// Mitsubishi GX Works2 project: 30国轩预化成10.29   PLC: Q10UDEH (continued)

Rotor30403(ShuttleCarInOut:=RotorIO30403);(*预化成2入库转台*)
RotorIO30403.xReady:=XAD;
Y264:=RotorIO30403.xCW;					
Y265:=RotorIO30403.xCCW;	
Y285:=RotorIO30403.xBrake;				
RotorIO30403.xForward:=M545;					
RotorIO30403.xBackward:=M546;					
ShuttleCarCurrentPosition(X65 OR X64,X65,X64,FALSE,RotorIO30403.iCurrentPos);					
M647:=RotorIO30403.xOvertimeAlarm ;					
RotorIO30403.diDeviceID:=30403;					
RotorIO30403.xPosLimit:=X6C;					
RotorIO30403.xNegLimit:=X6D;					

Rotor30404(ShuttleCarInOut:=RotorIO30404);(*预化成2出库转台*)
RotorIO30404.xReady:=XAE;
Y267:=RotorIO30404.xCW;					
Y266:=RotorIO30404.xCCW;	
Y286:=RotorIO30404.xBrake;					
RotorIO30404.xForward:=M547;					
RotorIO30404.xBackward:=M548;					
ShuttleCarCurrentPosition(X67 OR X66,X66,X67,FALSE,RotorIO30404.iCurrentPos);					
M648:=RotorIO30404.xOvertimeAlarm ;					
RotorIO30404.diDeviceID:=30404;					
RotorIO30404.xPosLimit:=X6E;					
RotorIO30404.xNegLimit:=X6F;					

Lifter30201(ShuttleCarInOut:=LifterIO30201);
LifterIO30201.xCylinder:=1;
Y22A:=LifterIO30201.xCW;					
Y22B:=LifterIO30201.xCCW;					
LifterIO30201.xForward:=M549;					
LifterIO30201.xBackward:=M550;					
ShuttleCarCurrentPosition(X2C OR X2B,X2C,X2B,FALSE,LifterIO30201.iCurrentPos);					
M649:=LifterIO30201.xOvertimeAlarm ;					
LifterIO30201.diDeviceID:=30201;					

Lifter30202(ShuttleCarInOut:=LifterIO30202);
LifterIO30202.xCylinder:=1;
Y22C:=LifterIO30202.xCW;					
Y22D:=LifterIO30202.xCCW;					
LifterIO30202.xForward:=M551;					
LifterIO30202.xBackward:=M552;					
ShuttleCarCurrentPosition(X2E OR X2D,X2E,X2D,FALSE,LifterIO30202.iCurrentPos);					
M650:=LifterIO30202.xOvertimeAlarm ;					
LifterIO30202.diDeviceID:=30202;					

Lifter30203(ShuttleCarInOut:=LifterIO30203);
LifterIO30203.xCylinder:=1;
Y22E:=LifterIO30203.xCW;					
Y22F:=LifterIO30203.xCCW;					
LifterIO30203.xForward:=M553;					
LifterIO30203.xBackward:=M554;					
ShuttleCarCurrentPosition(X30 OR X2F,X30,X2F,FALSE,LifterIO30203.iCurrentPos);					
M651:=LifterIO30203.xOvertimeAlarm ;					
LifterIO30203.diDeviceID:=30203;					

Lifter30204(ShuttleCarInOut:=LifterIO30204);
LifterIO30204.xCylinder:=1;
Y230:=LifterIO30204.xCW;					
Y231:=LifterIO30204.xCCW;					
LifterIO30204.xForward:=M555;					
LifterIO30204.xBackward:=M556;					
ShuttleCarCurrentPosition(X32 OR X31,X32,X31,FALSE,LifterIO30204.iCurrentPos);					
M652:=LifterIO30204.xOvertimeAlarm ;					
LifterIO30204.diDeviceID:=30204;					

Lifter30205(ShuttleCarInOut:=LifterIO30205);
LifterIO30205.xCylinder:=1;
Y232:=LifterIO30205.xCW;					
Y233:=LifterIO30205.xCCW;					
LifterIO30205.xForward:=M557;					
LifterIO30205.xBackward:=M558;					
ShuttleCarCurrentPosition(X34 OR X33,X34,X33,FALSE,LifterIO30205.iCurrentPos);					
M653:=LifterIO30205.xOvertimeAlarm ;					
LifterIO30205.diDeviceID:=30205;					

Lifter30206(ShuttleCarInOut:=LifterIO30206);
LifterIO30206.xCylinder:=1;
Y234:=LifterIO30206.xCW;					
Y235:=LifterIO30206.xCCW;					
LifterIO30206.xForward:=M559;					
LifterIO30206.xBackward:=M560;					
ShuttleCarCurrentPosition(X36 OR X35,X36,X35,FALSE,LifterIO30206.iCurrentPos);					
M654:=LifterIO30206.xOvertimeAlarm ;					
LifterIO30206.diDeviceID:=30206;					

Lifter30207(ShuttleCarInOut:=LifterIO30207);
LifterIO30207.xCylinder:=1;
Y238:=LifterIO30207.xCW;					
Y239:=LifterIO30207.xCCW;					
LifterIO30207.xForward:=M561;					
LifterIO30207.xBackward:=M562;					
ShuttleCarCurrentPosition(X3A OR X39,X3A,X39,FALSE,LifterIO30207.iCurrentPos);					
M655:=LifterIO30207.xOvertimeAlarm ;					
LifterIO30207.diDeviceID:=30207;					

Lifter30212(ShuttleCarInOut:=LifterIO30212);
LifterIO30212.xCylinder:=1;
Y254:=LifterIO30212.xCW;					
Y255:=LifterIO30212.xCCW;					
LifterIO30212.xForward:=M563;					
LifterIO30212.xBackward:=M564;					
ShuttleCarCurrentPosition(X58 OR X57,X57,X58,FALSE,LifterIO30212.iCurrentPos);					
M656:=LifterIO30212.xOvertimeAlarm ;					
LifterIO30212.diDeviceID:=30212;					

Lifter30213(ShuttleCarInOut:=LifterIO30213);
LifterIO30213.xCylinder:=1;
Y256:=LifterIO30213.xCW;					
Y257:=LifterIO30213.xCCW;					
LifterIO30213.xForward:=M565;					
LifterIO30213.xBackward:=M566;					
ShuttleCarCurrentPosition(X5A OR X59,X59,X5A,FALSE,LifterIO30213.iCurrentPos);					
M657:=LifterIO30213.xOvertimeAlarm ;					
LifterIO30213.diDeviceID:=30213;					

Lifter30214(ShuttleCarInOut:=LifterIO30214);(*预化成1出库末端顶起机构*)
LifterIO30214.xCylinder:=1;
Y258:=LifterIO30214.xCW;					
Y259:=LifterIO30214.xCCW;					
LifterIO30214.xForward:=M567;					
LifterIO30214.xBackward:=M568;					
ShuttleCarCurrentPosition(X5C OR X5B,X5B,X5C,FALSE,LifterIO30214.iCurrentPos);					
M658:=LifterIO30214.xOvertimeAlarm ;					
LifterIO30214.diDeviceID:=30214;					

Lifter30215(ShuttleCarInOut:=LifterIO30215);(*预化成1入库末端顶起机构*)
LifterIO30215.xCylinder:=1;
Y25A:=LifterIO30215.xCW;					
Y25B:=LifterIO30215.xCCW;					
LifterIO30215.xForward:=M569;					
LifterIO30215.xBackward:=M570;					
ShuttleCarCurrentPosition(X5E OR X5D,X5D,X5E,FALSE,LifterIO30215.iCurrentPos);					
M659:=LifterIO30215.xOvertimeAlarm ;					
LifterIO30215.diDeviceID:=30215;					

Switch30301(ConveyorEntryIO:=ConveyorIO30101 ,ConveyorExitIO:=ConveyorIO30102 ,SwitchIO:=SwitchIO30301);
SwitchIO30301.xLiftCylinderRetractDetect:=X3E;							
SwitchIO30301.xLiftCylinderExtendDetect:=X3D;							
Y23A:=SwitchIO30301.xLiftCylinderExtend;							
SwitchIO30301.xLiftCylinderExtendButton:=M571;	
SwitchIO30301.xLiftCylinderRetractButton:=NOT M571;
(*阻挡气缸暂时没接*)(*装了死挡*)
Y288:=NOT SwitchIO30301.xExitBarCylinderRetract;						
M660:=SwitchIO30301.xOvertimeAlarm ;							

Switch30302(ConveyorEntryIO:=ConveyorIO30103 ,ConveyorExitIO:=ConveyorIO30141 ,SwitchIO:=SwitchIO30302);
SwitchIO30302.xLiftCylinderExtendInit:=1;
SwitchIO30302.xLiftCylinderRetractDetect:=X40;							
SwitchIO30302.xLiftCylinderExtendDetect:=X3F;							
Y23C:=SwitchIO30302.xLiftCylinderExtend;							
SwitchIO30302.xLiftCylinderExtendButton:=M572;	
SwitchIO30302.xLiftCylinderRetractButton:=NOT M572;						
M661:=SwitchIO30302.xOvertimeAlarm ;							

Switch30303(ConveyorEntryIO:=ConveyorIO30107 ,ConveyorExitIO:=ConveyorIO30105 ,SwitchIO:=SwitchIO30303);
SwitchIO30303.xLiftCylinderExtendInit:=1;
SwitchIO30303.xLiftCylinderRetractDetect:=X42;							
SwitchIO30303.xLiftCylinderExtendDetect:=X41;							
Y23E:=SwitchIO30303.xLiftCylinderExtend;							
SwitchIO30303.xLiftCylinderExtendButton:=M573;	
SwitchIO30303.xLiftCylinderRetractButton:=NOT M573;						
M662:=SwitchIO30303.xOvertimeAlarm ;							

Switch30304(ConveyorEntryIO:=ConveyorIO30142 ,ConveyorExitIO:=ConveyorIO30108 ,SwitchIO:=SwitchIO30304);
SwitchIO30304.xLiftCylinderRetractDetect:=X44;							
SwitchIO30304.xLiftCylinderExtendDetect:=X43;							
Y240:=SwitchIO30304.xLiftCylinderExtend;							
SwitchIO30304.xLiftCylinderExtendButton:=M574;	
SwitchIO30304.xLiftCylinderRetractButton:=NOT M574;
M663:=SwitchIO30304.xOvertimeAlarm ;							

Switch30305(ConveyorEntryIO:=ConveyorIO30106 ,ConveyorExitIO:=ConveyorIO30111 ,SwitchIO:=SwitchIO30305);
SwitchIO30305.xLiftCylinderRetractDetect:=X46;							
SwitchIO30305.xLiftCylinderExtendDetect:=X45;							
Y242:=SwitchIO30305.xLiftCylinderExtend;							
Y28A:=SwitchIO30305.xExitBarCylinderRetract;							
SwitchIO30305.xLiftCylinderExtendButton:=M575;	
SwitchIO30305.xLiftCylinderRetractButton:=NOT M575;						
SwitchIO30305.xExitBarCylinderRetractButton:=M576;							
M664:=SwitchIO30305.xOvertimeAlarm ;							

Switch30306(ConveyorEntryIO:=ConveyorIO30113 ,ConveyorExitIO:=ConveyorIO30110 ,SwitchIO:=SwitchIO30306);
SwitchIO30306.xLiftCylinderExtendInit:=1;
SwitchIO30306.xLiftCylinderRetractDetect:=X47;							
SwitchIO30306.xLiftCylinderExtendDetect:=X48;							
Y244:=SwitchIO30306.xLiftCylinderExtend;							
SwitchIO30306.xLiftCylinderExtendButton:=M577;	
SwitchIO30306.xLiftCylinderRetractButton:=NOT M577;						
M665:=SwitchIO30306.xOvertimeAlarm ;							

Switch30307(ConveyorEntryIO:=ConveyorIO30115 ,ConveyorExitIO:=ConveyorIO30116 ,SwitchIO:=SwitchIO30307);
SwitchIO30307.xLiftCylinderRetractDetect:=X4A;							
SwitchIO30307.xLiftCylinderExtendDetect:=X49;							
Y246:=SwitchIO30307.xLiftCylinderExtend;							
Y28C:=SwitchIO30307.xExitBarCylinderRetract;							
SwitchIO30307.xLiftCylinderExtendButton:=M578;	
SwitchIO30307.xLiftCylinderRetractButton:=NOT M578;						
SwitchIO30307.xExitBarCylinderRetractButton:=M579;							
M666:=SwitchIO30307.xOvertimeAlarm ;							

Switch30308(ConveyorEntryIO:=ConveyorIO30118 ,ConveyorExitIO:=ConveyorIO30122 ,SwitchIO:=SwitchIO30308);
SwitchIO30308.xLiftCylinderExtendInit:=1;
SwitchIO30308.xLiftCylinderRetractDetect:=X4B;							
SwitchIO30308.xLiftCylinderExtendDetect:=X4C;							
Y248:=SwitchIO30308.xLiftCylinderExtend;							
SwitchIO30308.xLiftCylinderExtendButton:=M580;
SwitchIO30308.xLiftCylinderRetractButton:=NOT M580;
M667:=SwitchIO30308.xOvertimeAlarm ;							

Switch30309(ConveyorEntryIO:=ConveyorIO30126 ,ConveyorExitIO:=ConveyorIO30127 ,SwitchIO:=SwitchIO30309);
SwitchIO30309.xLiftCylinderRetractDetect:=X52;							
SwitchIO30309.xLiftCylinderExtendDetect:=X51;							
Y24E:=SwitchIO30309.xLiftCylinderExtend;							
Y293:=SwitchIO30309.xExitBarCylinderRetract;							
SwitchIO30309.xLiftCylinderExtendButton:=M581;							
SwitchIO30309.xExitBarCylinderRetractButton:=M582;							
M668:=SwitchIO30309.xOvertimeAlarm ;							

Switch30310(ConveyorEntryIO:=ConveyorIO301271 ,ConveyorExitIO:=ConveyorIO30128 ,SwitchIO:=SwitchIO30310);
SwitchIO30310.xLiftCylinderExtendInit:=1;
SwitchIO30310.xLiftCylinderRetractDetect:=X54;							
SwitchIO30310.xLiftCylinderExtendDetect:=X53;							
Y250:=SwitchIO30310.xLiftCylinderExtend;							
SwitchIO30310.xLiftCylinderExtendButton:=M583;							
M669:=SwitchIO30310.xOvertimeAlarm ;							

Switch30311(ConveyorEntryIO:=ConveyorIO30139 ,ConveyorExitIO:=ConveyorIO301201 ,SwitchIO:=SwitchIO30311);
SwitchIO30311.xLiftCylinderRetractDetect:=X56;							
SwitchIO30311.xLiftCylinderExtendDetect:=X55;							
Y252:=SwitchIO30311.xLiftCylinderExtend;							
Y291:=SwitchIO30311.xExitBarCylinderRetract;							
SwitchIO30311.xLiftCylinderExtendButton:=M584;							
SwitchIO30311.xExitBarCylinderRetractButton:=M585;							
M670:=SwitchIO30311.xOvertimeAlarm ;							
(****************上位机通信数据************************)
(*24H入库扫码*)
ComConveyor30103(ConveyorIO:=ConveyorIO301021,CommunicationIO:=ComConveyorIO30103);
ComConveyorIO30103.i_iResponsPCPLC:=D2000;	
ComConveyorIO30103.i_iTypeInfoPCPLC:=D2001;
ComConveyorIO30103.i_iReadWriteFlagPCPLC:=D2005;	
ComConveyorIO30103.i_iTaskProcessFlagPCPLC:=D2006;	
ComConveyorIO30103.i_iCommandPCPLC:=D2007;	
ComConveyorIO30103.i_iTaskIDPCPLC:=D2008;	
DMOV(TRUE,D2009,ComConveyorIO30103.i_diDestinationDevicePCPLC);	
ComConveyorIO30103.i_iProductIDPCPLC:=D2011;	
D3000:=ComConveyorIO30103.o_iRequestPLCPC;	
D3001:=ComConveyorIO30103.o_iForceInportPLCPC;
D3002:=ComConveyorIO30103.o_iFolderNumberPLCPC;
D3003:=ComConveyorIO30103.o_iEmptyPLCPC;
D3005:=ComConveyorIO30103.o_iReadWriteFlagPLCPC;	
D3006:=ComConveyorIO30103.o_iDeviceStatusPLCPC;	
D3007:=ComConveyorIO30103.o_iTaskIDPLCPC;	
D3008:=ComConveyorIO30103.o_iProductIDPLCPC;	
(*入库站台1*)
ComConveyor30136(ConveyorIO:=ConveyorIO30136,CommunicationIO:=ComConveyorIO30136);
ComConveyorIO30136.i_iResponsPCPLC:=D2015;	
ComConveyorIO30136.i_iTypeInfoPCPLC:=D2016;
ComConveyorIO30136.i_iReadWriteFlagPCPLC:=D2020;	
ComConveyorIO30136.i_iTaskProcessFlagPCPLC:=D2021;	
ComConveyorIO30136.i_iCommandPCPLC:=D2022;	
ComConveyorIO30136.i_iTaskIDPCPLC:=D2023;	
DMOV(TRUE,D2024,ComConveyorIO30136.i_diDestinationDevicePCPLC);	
ComConveyorIO30136.i_iProductIDPCPLC:=D2026;	
D3015:=ComConveyorIO30136.o_iRequestPLCPC;	
D3016:=ComConveyorIO30136.o_iForceInportPLCPC;
D3017:=ComConveyorIO30136.o_iFolderNumberPLCPC;
D3018:=ComConveyorIO30136.o_iEmptyPLCPC;
D3020:=ComConveyorIO30136.o_iReadWriteFlagPLCPC;	
D3021:=ComConveyorIO30136.o_iDeviceStatusPLCPC;	
D3022:=ComConveyorIO30136.o_iTaskIDPLCPC;	
D3023:=ComConveyorIO30136.o_iProductIDPLCPC;	
ComConveyorIO30136.i_xExtraCondition:=NOT g_x24HourImport1Forbidden;(*触摸屏上的按钮，重新提交任务*)
(*入库站台2*)
ComConveyor30104(ConveyorIO:=ConveyorIO30104,CommunicationIO:=ComConveyorIO30104);
ComConveyorIO30104.i_iResponsPCPLC:=D2030;	
ComConveyorIO30104.i_iTypeInfoPCPLC:=D2031;
ComConveyorIO30104.i_iReadWriteFlagPCPLC:=D2035;	
ComConveyorIO30104.i_iTaskProcessFlagPCPLC:=D2036;	
ComConveyorIO30104.i_iCommandPCPLC:=D2037;	
ComConveyorIO30104.i_iTaskIDPCPLC:=D2038;	
DMOV(TRUE,D2039,ComConveyorIO30104.i_diDestinationDevicePCPLC);	
ComConveyorIO30104.i_iProductIDPCPLC:=D2041;	
D3030:=ComConveyorIO30104.o_iRequestPLCPC;	
D3031:=ComConveyorIO30104.o_iForceInportPLCPC;
D3032:=ComConveyorIO30104.o_iFolderNumberPLCPC;
D3033:=ComConveyorIO30104.o_iEmptyPLCPC;
D3035:=ComConveyorIO30104.o_iReadWriteFlagPLCPC;	
D3036:=ComConveyorIO30104.o_iDeviceStatusPLCPC;	
D3037:=ComConveyorIO30104.o_iTaskIDPLCPC;	
D3038:=ComConveyorIO30104.o_iProductIDPLCPC;	
ComConveyorIO30104.i_xExtraCondition:=NOT g_x24HourImport2Forbidden;(*触摸屏上的按钮，重新提交任务*)
(*出库站台1*)
ComConveyor30137(ConveyorIO:=ConveyorIO30137,CommunicationIO:=ComConveyorIO30137);
ComConveyorIO30137.i_iResponsPCPLC:=D2045;	
ComConveyorIO30137.i_iTypeInfoPCPLC:=D2046;
ComConveyorIO30137.i_iReadWriteFlagPCPLC:=D2050;	
ComConveyorIO30137.i_iTaskProcessFlagPCPLC:=D2051;	
ComConveyorIO30137.i_iCommandPCPLC:=D2052;	
ComConveyorIO30137.i_iTaskIDPCPLC:=D2053;	
DMOV(TRUE,D2054,ComConveyorIO30137.i_diDestinationDevicePCPLC);	
ComConveyorIO30137.i_iProductIDPCPLC:=D2056;	
D3045:=ComConveyorIO30137.o_iRequestPLCPC;	
D3046:=ComConveyorIO30137.o_iForceInportPLCPC;
D3047:=ComConveyorIO30137.o_iFolderNumberPLCPC;
D3048:=ComConveyorIO30137.o_iEmptyPLCPC;
D3050:=ComConveyorIO30137.o_iReadWriteFlagPLCPC;	
D3051:=ComConveyorIO30137.o_iDeviceStatusPLCPC;	
D3052:=ComConveyorIO30137.o_iTaskIDPLCPC;	
D3053:=ComConveyorIO30137.o_iProductIDPLCPC;	
ComConveyorIO30137.i_xExtraCondition:=ConveyorIO30109.xEmpty AND NOT ConveyorIO30109.xCWPresent  AND NOT ConveyorIO30137.xCWPresent 
																						AND NOT g_x24HourExport1Forbidden;(*无出库禁止*)
ComConveyorIO30137.i_xExportConveyor:=1;
(*预化成1入库转台前扫码*)
ComConveyor30111(ConveyorIO:=ConveyorIO30134,CommunicationIO:=ComConveyorIO30111);
ComConveyorIO30111.i_iResponsPCPLC:=D2060;	
ComConveyorIO30111.i_iTypeInfoPCPLC:=D2061;
ComConveyorIO30111.i_iReadWriteFlagPCPLC:=D2065;	
ComConveyorIO30111.i_iTaskProcessFlagPCPLC:=D2066;	
ComConveyorIO30111.i_iCommandPCPLC:=D2067;	
ComConveyorIO30111.i_iTaskIDPCPLC:=D2068;	
DMOV(TRUE,D2069,ComConveyorIO30111.i_diDestinationDevicePCPLC);	
ComConveyorIO30111.i_iProductIDPCPLC:=D2071;	
D3060:=ComConveyorIO30111.o_iRequestPLCPC;	
D3061:=ComConveyorIO30111.o_iForceInportPLCPC;
D3062:=ComConveyorIO30111.o_iFolderNumberPLCPC;
D3063:=ComConveyorIO30111.o_iEmptyPLCPC;
D3065:=ComConveyorIO30111.o_iReadWriteFlagPLCPC;	
D3066:=ComConveyorIO30111.o_iDeviceStatusPLCPC;	
D3067:=ComConveyorIO30111.o_iTaskIDPLCPC;	
D3068:=ComConveyorIO30111.o_iProductIDPLCPC;	
ComConveyorIO30111.i_xExtraCondition:=ConveyorIO30112.xEmpty AND NOT ConveyorIO30112.xCWPresent  (*入库这里确定后面无料再发扫码请求*)
																						 AND lifterio30215.iCurrentPos=1 AND X5D;    (*还要判断顶升位置，因为没装漫反射,可能出现误判断*)
(*预化成2入库转台扫码*)
ComConveyor30116(ConveyorIO:=ConveyorIO30132,CommunicationIO:=ComConveyorIO30116);
ComConveyorIO30116.i_iResponsPCPLC:=D207(*5*);	
ComConveyorIO30116.i_iTypeInfoPCPLC:=D2076;
ComConveyorIO30116.i_iReadWriteFlagPCPLC:=D2080;	
ComConveyorIO30116.i_iTaskProcessFlagPCPLC:=D2081;	
ComConveyorIO30116.i_iCommandPCPLC:=D2082;	
ComConveyorIO30116.i_iTaskIDPCPLC:=D2083;	
DMOV(TRUE,D2084,ComConveyorIO30116.i_diDestinationDevicePCPLC);	
ComConveyorIO30116.i_iProductIDPCPLC:=D2086;	
D3075:=ComConveyorIO30116.o_iRequestPLCPC;	
D3076:=ComConveyorIO30116.o_iForceInportPLCPC;
D3077:=ComConveyorIO30116.o_iFolderNumberPLCPC;
D3078:=ComConveyorIO30116.o_iEmptyPLCPC;
D3080:=ComConveyorIO30116.o_iReadWriteFlagPLCPC;	
D3081:=ComConveyorIO30116.o_iDeviceStatusPLCPC;	
D3082:=ComConveyorIO30116.o_iTaskIDPLCPC;	
D3083:=ComConveyorIO30116.o_iProductIDPLCPC;	
ComConveyorIO30116.i_xExtraCondition:=ConveyorIO30117.xEmpty AND NOT ConveyorIO30117.xCWPresent  (*入库这里确定后面无料再发扫码请求*)
																						 AND lifterio30213.iCurrentPos=1 AND X59;    (*还要判断顶升位置，因为没装漫反射,可能出现误判断*)

(*化成1入库站台*)
ComConveyor30112(ConveyorIO:=ConveyorIO30112,CommunicationIO:=ComConveyorIO30112);
ComConveyorIO30112.i_iResponsPCPLC:=D2090;	
ComConveyorIO30112.i_iTypeInfoPCPLC:=D2091;
ComConveyorIO30112.i_iReadWriteFlagPCPLC:=D2095;	
ComConveyorIO30112.i_iTaskProcessFlagPCPLC:=D2096;	
ComConveyorIO30112.i_iCommandPCPLC:=D2097;	
ComConveyorIO30112.i_iTaskIDPCPLC:=D2098;	
DMOV(TRUE,D2099,ComConveyorIO30112.i_diDestinationDevicePCPLC);	
ComConveyorIO30112.i_iProductIDPCPLC:=D2101;	
D3090:=ComConveyorIO30112.o_iRequestPLCPC;	
D3091:=ComConveyorIO30112.o_iForceInportPLCPC;
D3092:=ComConveyorIO30112.o_iFolderNumberPLCPC;
D3093:=ComConveyorIO30112.o_iEmptyPLCPC;
D3095:=ComConveyorIO30112.o_iReadWriteFlagPLCPC;	
D3096:=ComConveyorIO30112.o_iDeviceStatusPLCPC;	
D3097:=ComConveyorIO30112.o_iTaskIDPLCPC;	
D3098:=ComConveyorIO30112.o_iProductIDPLCPC;	
ComConveyorIO30112.i_xExtraCondition:=LifterIO30215.iCurrentPos=2 
																					AND NOT g_xPreChemImport1Forbidden;(*且没有入库禁止，禁止了就不报完成，就不生成任务了*)
(*这里加一个条件，当位置在2时，不在触摸屏上显示禁止按钮*)

(*化成2入库站台*)
ComConveyor30117(ConveyorIO:=ConveyorIO30117,CommunicationIO:=ComConveyorIO30117);
ComConveyorIO30117.i_iResponsPCPLC:=D2105;	
ComConveyorIO30117.i_iTypeInfoPCPLC:=D2106;
ComConveyorIO30117.i_iReadWriteFlagPCPLC:=D2110;	
ComConveyorIO30117.i_iTaskProcessFlagPCPLC:=D2111;	
ComConveyorIO30117.i_iCommandPCPLC:=D2112;	
ComConveyorIO30117.i_iTaskIDPCPLC:=D2113;	
DMOV(TRUE,D2114,ComConveyorIO30117.i_diDestinationDevicePCPLC);	
ComConveyorIO30117.i_iProductIDPCPLC:=D2116;	
D3105:=ComConveyorIO30117.o_iRequestPLCPC;	
D3106:=ComConveyorIO30117.o_iForceInportPLCPC;
D3107:=ComConveyorIO30117.o_iFolderNumberPLCPC;
D3108:=ComConveyorIO30117.o_iEmptyPLCPC;
D3110:=ComConveyorIO30117.o_iReadWriteFlagPLCPC;	
D3111:=ComConveyorIO30117.o_iDeviceStatusPLCPC;	
D3112:=ComConveyorIO30117.o_iTaskIDPLCPC;	
D3113:=ComConveyorIO30117.o_iProductIDPLCPC;	
ComConveyorIO30117.i_xExtraCondition:=LifterIO30213.iCurrentPos=2
																				AND NOT g_xPreChemImport2Forbidden;(*且没有入库禁止，禁止了就不扫码*)

(*化成1出库站台*)
ComConveyor30114(ConveyorIO:=ConveyorIO30114,CommunicationIO:=ComConveyorIO30114);
ComConveyorIO30114.i_iResponsPCPLC:=D2120;	
ComConveyorIO30114.i_iTypeInfoPCPLC:=D2121;
ComConveyorIO30114.i_iReadWriteFlagPCPLC:=D2125;	
ComConveyorIO30114.i_iTaskProcessFlagPCPLC:=D2126;	
ComConveyorIO30114.i_iCommandPCPLC:=D2127;	
ComConveyorIO30114.i_iTaskIDPCPLC:=D2128;	
DMOV(TRUE,D2129,ComConveyorIO30114.i_diDestinationDevicePCPLC);	
ComConveyorIO30114.i_iProductIDPCPLC:=D2131;	
D3120:=ComConveyorIO30114.o_iRequestPLCPC;	
D3121:=ComConveyorIO30114.o_iForceInportPLCPC;
D3122:=ComConveyorIO30114.o_iFolderNumberPLCPC;
D3123:=ComConveyorIO30114.o_iEmptyPLCPC;
D3125:=ComConveyorIO30114.o_iReadWriteFlagPLCPC;	
D3126:=ComConveyorIO30114.o_iDeviceStatusPLCPC;	
D3127:=ComConveyorIO30114.o_iTaskIDPLCPC;	
D3128:=ComConveyorIO30114.o_iProductIDPLCPC;	
ComConveyorIO30114.i_xExportConveyor:=1;
ComConveyorIO30114.i_xExtraCondition:=NOT ConveyorIO30114.xCCWPresent AND LifterIO30214.iCurrentPos=2 
																					AND ConveyorIO30133.xEmpty AND NOT ConveyorIO30133.xCWPresent
																					AND NOT g_xPreChemExport1Forbidden;
(*化成2出库站台*)
ComConveyor30119(ConveyorIO:=ConveyorIO30119,CommunicationIO:=ComConveyorIO30119);
ComConveyorIO30119.i_iResponsPCPLC:=D2135;	
ComConveyorIO30119.i_iTypeInfoPCPLC:=D2136;
ComConveyorIO30119.i_iReadWriteFlagPCPLC:=D2140;	
ComConveyorIO30119.i_iTaskProcessFlagPCPLC:=D2141;	
ComConveyorIO30119.i_iCommandPCPLC:=D2142;	
ComConveyorIO30119.i_iTaskIDPCPLC:=D2143;	
DMOV(TRUE,D2144,ComConveyorIO30119.i_diDestinationDevicePCPLC);	
ComConveyorIO30119.i_iProductIDPCPLC:=D2146;	
D3135:=ComConveyorIO30119.o_iRequestPLCPC;	
D3136:=ComConveyorIO30119.o_iForceInportPLCPC;
D3137:=ComConveyorIO30119.o_iFolderNumberPLCPC;
D3138:=ComConveyorIO30119.o_iEmptyPLCPC;
D3140:=ComConveyorIO30119.o_iReadWriteFlagPLCPC;	
D3141:=ComConveyorIO30119.o_iDeviceStatusPLCPC;	
D3142:=ComConveyorIO30119.o_iTaskIDPLCPC;	
D3143:=ComConveyorIO30119.o_iProductIDPLCPC;	
ComConveyorIO30119.i_xExportConveyor:=1;
ComConveyorIO30119.i_xExtraCondition:=NOT ConveyorIO30119.xCCWPresent AND LifterIO30212.iCurrentPos=2 
																					AND ConveyorIO30131.xEmpty AND NOT ConveyorIO30131.xCWPresent
																					AND NOT g_xPreChemExport2Forbidden;
(*不良品分拣工位*)

SortConveyor30121(ConveyorIO:=ConveyorIO30121 ,SortCommunicationIO:= SortConveyorIO30121 ,FanucRobotIO:=FanucRobotIO300);
SortConveyorIO30121 .i_iResponsPCPLC:=D2240;
SortConveyorIO30121 .i_iInfoWriteDone:=D2241;
SortConveyorIO30121 .i_iSortDoneAknPCPLC:=D2242;
D3240:=SortConveyorIO30121 .o_iRequestPLCPC;(*有料请求*)
D3241:=SortConveyorIO30121 .o_iSortDonePLCPC;(*分拣完成信号*)
FOR Z0:=0 TO 127 BY 1 DO
	SortConveyorIO30121 .i_arriBatteryStatus[Z0+1]:=D2243Z0;
END_FOR;

(****************以上是上位机通信数据************************)
(**********以下是自动程序***************************************)
IF g_xAuto THEN
(*高温静置库上料*)
	D201.2:=ConveyorIO30101.xEmpty;
	SwitchIO30301.xEntryEnable:=D401.2 OR M8;
	SwitchIO30301.xSwithEnable:=1;
	SwitchIO30301.xExitEnable:=(*LifterIO30202.iCurrentPos=2 AND*) ConveyorIO301021.xEmpty;(*等门升起再下料*)
(*门的升降控制*)	
	IF ConveyorIO301021.xEmpty AND NOT ConveyorIO30102.xEmpty THEN
		LifterIO30201.xMDIExe:=1;
		LifterIO30201.iDestinationPos:=2;
	ELSIF NOT	ConveyorIO301021.xEmpty AND ConveyorIO30102.xEmpty 
				AND NOT ConveyorIO30102.xCWPresent THEN(*这里加个开关的限制，防止直接下降压到电池*)
		LifterIO30201.xMDIExe:=1;
		LifterIO30201.iDestinationPos:=1;
	END_IF;	
(*运到待料站台*)
 	ConveyorIO301021.xLoad:=ConveyorIO30102.xNextRun;
 	ConveyorIO301021.xUnload:=ConveyorIO30103.xEmpty 
 															AND ConveyorIO301021.diDesConveyor<>0;
	(*数据传递,021传给03,03通过switch给到41，41给04,04给36*)
 	ConveyorIO30103.diDesConveyorIn:=ConveyorIO301021.diDesConveyorOut;
 	ConveyorIO30103.iProductCategoryIn:=ConveyorIO301021.iProductCategoryOut;
 	ConveyorIO30103.iTaskIDIn:=ConveyorIO301021.iTaskIDOut;
 	ConveyorIO30104.diDesConveyorIn:=ConveyorIO30141.diDesConveyorOut;
 	ConveyorIO30104.iProductCategoryIn:=ConveyorIO30141.iProductCategoryOut;
 	ConveyorIO30104.iTaskIDIn:=ConveyorIO30141.iTaskIDOut; 
 	 ConveyorIO30136.diDesConveyorIn:=ConveyorIO30104.diDesConveyorOut;
 	ConveyorIO30136.iProductCategoryIn:=ConveyorIO30104.iProductCategoryOut;
 	ConveyorIO30136.iTaskIDIn:=ConveyorIO30104.iTaskIDOut;
 	(*物料输送*)
 	SwitchIO30302.xEntryEnable:=ConveyorIO301021.xNextRun;
	SwitchIO30302.xSwithEnable:=1;
	SwitchIO30302.xExitEnable:=ConveyorIO30104.xEmpty(*肯定要等104为空*)
														AND(ConveyorIO30103.diDesConveyor=30104 (*目标104就不判断136状态*)
																	OR ConveyorIO30103.diDesConveyor=30136 AND ConveyorIO30136.xEmpty)  ;(*如果目标136，就需要136为空*)
	ConveyorIO30104.xLoad:=ConveyorIO30141.xNextRun;
	ConveyorIO30104.xUnload:=ConveyorIO30136.xEmpty AND ConveyorIO30104.diDesConveyor=30136;
	ConveyorIO30136.xLoad:=ConveyorIO30104.xNextRun;

	
	
	(*两段线体的putinto信号在通信块里写好了，所以这里就不写了。*)
	(*暂时这么写，有上位机再屏蔽*)
	SET(LDP(TRUE, NOT ConveyorIO30104.xBusy AND SM412),ConveyorIO30104.xPutInto);
	RST(LDF(TRUE, NOT ConveyorIO30104.xBusy AND SM412),ConveyorIO30104.xPutInto);
	SET(LDP(TRUE, NOT ConveyorIO30104.xBusy AND SM412),ConveyorIO30136.xPutInto);
	RST(LDF(TRUE,NOT  ConveyorIO30104.xBusy AND SM412),ConveyorIO30136.xPutInto);
(*针对下面这种情况，就需要能自动复位*)
	IF LDP(TRUE, NOT ConveyorIO30103.xEmpty AND NOT ConveyorIO30103.xCWPresent AND NOT ConveyorIO30141.xBusy) THEN
		ConveyorIO30103.xPutInto:=1;(*有料却没感应到开关，就不对劲，刷掉*)
	ELSIF 	ConveyorIO30103.xEmpty THEN
		ConveyorIO30103.xPutInto:=0;
END_IF;
	(*如果连续两筐都是一个地址，这时候会卡，所以需要强制入库*)	
	IF (ConveyorIO30103.diDesConveyor=30136 AND NOT ConveyorIO30136.xEmpty
																							AND NOT ConveyorIO30103.xEmpty AND ConveyorIO30103.xCWPresent(*加一个开关限制，防止开关误动作导致错误*)
																							AND ConveyorIO30104.xEmpty)
		OR g_xForceImport		THEN
		 ComConveyorIO30136.o_iForceInportPLCPC:=2;
		 ComConveyorIO30136.o_iRequestPLCPC:=2;
	ELSE
		 ComConveyorIO30136.o_iForceInportPLCPC:=1;
	END_IF;
	IF ConveyorIO30104.xEmpty AND ConveyorIO30136.xEmpty THEN
		g_xForceImport:=0;
	END_IF;	
	(*
	ConveyorIO30137.xPutInto:=NOT ConveyorIO30137.xBusy AND SM413;*)
(********************************高温库出库********************)	
	(*出库线体只有末端有通信，前面那段没通信，所以需要程序里给putinto信号*)
	ConveyorIO30109.xPutInto:=ConveyorIO30137.xPutInto;
	ConveyorIO30137.xUnload:=ConveyorIO30109.xEmpty;
	ConveyorIO30109.xLoad:=ConveyorIO30137.xNextRun;
	ConveyorIO30109.xUnload:=ConveyorIO30142.xEmpty;
	SwitchIO30304.xEntryEnable:=ConveyorIO30109.xNextRun;
	SwitchIO30304.xSwithEnable:=1;
	SwitchIO30304.xExitEnable:=ConveyorIO301071.xEmpty;
	ConveyorIO301071.xLoad:=ConveyorIO30108.xNextRun;
	ConveyorIO301071.xUnload:=ConveyorIO30107.xEmpty (* AND LifterIO30202.iCurrentPos=2*);
(*门的升降控制*)	
	IF ConveyorIO30107.xEmpty AND NOT ConveyorIO301071.xEmpty THEN
		LifterIO30202.xMDIExe:=1;
		LifterIO30202.iDestinationPos:=2;
	ELSIF NOT	ConveyorIO30107.xEmpty AND ConveyorIO301071.xEmpty 
				AND NOT ConveyorIO301071.xCWPresent THEN(*这里加个开关的限制，防止直接下降压到电池*)
		LifterIO30202.xMDIExe:=1;
		LifterIO30202.iDestinationPos:=1;
	END_IF;
(*静置库出库顶升移载*)		
	SwitchIO30303.xEntryEnable:=ConveyorIO301071.xNextRun;
	SwitchIO30303.xSwithEnable:=1;
	SwitchIO30303.xExitEnable:=ConveyorIO301051.xEmpty;
	ConveyorIO301051.xLoad:=ConveyorIO30105.xNextRun;
	ConveyorIO301051.xUnload:=ConveyorIO30106.xEmpty
						AND (m_iTask30303=2 (*2巷道任务*)
									OR (m_iTask30303=1 AND m_iTask30305=2));(*或1巷道但是是正常入库(305为2是正常入库,1是品检入库)*)
(***********************预化成12巷道的任务分配，排队任务，决定去哪个巷道*********************)	
	Task30303(arrxCondition:=Task30303Condition,
						xTaskComplete:= LDP(TRUE,ConveyorIO30106.xEmpty) ,
	 					xReset:=g_xResetSingle AND g_diDeviceIDSelect=30105 ,
						 iPriority:=m_iTask30303);
		Task30303Condition[1].xCondition :=m_xLocation1Empty  AND g_xLoadPermit[1];(*1巷道为空*)
		Task30303Condition[2].xCondition:= m_xLocation2Empty AND g_xLoadPermit[2];(*2巷道为空*)
		g_xLoadPermit[1]:=M50;(*任务可以通过触摸屏控制生成*)
		g_xLoadPermit[2]:=M51;
		DMOV(m_iTask30303=1,30112,ConveyorIO301051.diDesConveyor);(*30112是入库对接那段线体的ID*)
		DMOV(m_iTask30303=1,30112,ConveyorIO30106.diDesConveyor);(*是品检回流入库时，直接putinto的，就没有传递了，所以可以强制*)
		DMOV(m_iTask30303=2,30116,ConveyorIO301051.diDesConveyor);(*【初始目标地址的生成】*)
	(*以上是12巷道任务分配的排队任务*)	
(***********************1巷道入库的抢占任务，一边是正常分流入库，一边是品捡后回库*********************)	
	Task30305(xCondition:= Task30305Condition,(*抢栈式*)
						xTaskComplete:= LDP(TRUE,ConveyorIO30106.xEmpty),
	 					xReset:=g_xResetSingle AND g_diDeviceIDSelect=30106,
						 iPriority:=m_iTask30305);
		Task30305Condition[1]:=NOT ConveyorIO30140.xEmpty AND m_iTask30303=1 ;(*品检回流*)
		Task30305Condition[2]:=NOT ConveyorIO301051.xEmpty AND m_iTask30303=1  ;(*正常入库*)
	(*以上是1巷道的抢占任务*)	

	SwitchIO30305.xEntryEnable:=ConveyorIO301051.xNextRun;
	ConveyorIO30106.diDesConveyorIn:=ConveyorIO301051.diDesConveyorOut;(*【目标地址从1051传到106】*)
	SwitchIO30305.xSwithEnable:=ConveyorIO30106.diDesConveyor=30112;(*根据目标地址定是否转向，1巷道转，2巷道不转*)
	SwitchIO30305.xExitEnable:=(SwitchIO30305.xSwithEnable AND m_xLocation1Empty)(*需要转到1库，则1这边空就下料*)
															OR (NOT SwitchIO30305.xSwithEnable 
																	AND m_iTask30306=2 AND ConveyorIO30110.xEmpty(*不需要转，则等顶升移载306生成2任务*)
																	AND ConveyorIO30138.xEmpty);(*这里是因为10和38共用一个电机，所以必须都为empty才行*)
	IF m_iTask30303=1 AND m_iTask30305=1 THEN(*回流入库*)
		ConveyorIO30140.xUnload:=ConveyorIO30111.xEmpty;
		IF ConveyorIO30111.xEmpty THEN
			SwitchIO30305.xLiftCylinderExtend:=1;
			SwitchIO30305.xLiftCylinderRetract:=0;
		END_IF;
		ConveyorIO30111.xLoad:=ConveyorIO30140.xNextRun;(*这里运到11上，等待扫码，旋转，再往后运*)
		SET(LDP(TRUE,NOT ConveyorIO30111.xEmpty),ConveyorIO30106.xPutInto);(*这里只要putinto了，就会进入switch正常流程了*)
		RST(LDP(TRUE,NOT ConveyorIO30106.xEmpty),ConveyorIO30106.xPutInto);
	END_IF;
	m_xLocation1Load:=ConveyorIO30111.xNextRun;
(**************************************1巷道旋转，入库处理*****************************************************)
	(*定位机发出料请求，我要把门升起来，再给他发下料信号*)
	LifterIO30203.xMDIExe:=NOT ConveyorIO30134.xError;
		IF m_xLocation1NextRun AND ConveyorIO30134.xEmpty THEN
			LifterIO30203.iDestinationPos:=2;
		ELSE 
			LifterIO30203.iDestinationPos:=1;
		END_IF;	
	(*预化成1入库转台上料*)		
		m_xLocation1Unload:= ConveyorIO30134.xEmpty AND m_xLocation1NextRun(*他有下料请求时，我才判断*)
														AND RotorIO30401.iCurrentPos=1 AND X60(*转台在位置1才上料*)
														(*AND  LifterIO30203.iCurrentPos=2 AND X30*);												
		ConveyorIO30134.xLoad:=m_xLocation1NextRun 
															 AND RotorIO30401.iCurrentPos=1 AND X60
															(*AND  LifterIO30203.iCurrentPos=2 AND X30*) ;
	(*预化成1入库旋转控制*)		
		RotorIO30401.xMDIExe:=NOT ConveyorIO301111.xError AND NOT ConveyorIO30134.xError AND NOT ConveyorIO30112.xError;
	
			IF NOT ConveyorIO30134.xEmpty THEN(*有料时，旋转，转到2旋转完成*)
				ConveyorIO30134.xUnloadCCW:=ComConveyorIO30111.i_iResponsPCPLC=4;
				MOV(ComConveyorIO30111.i_iResponsPCPLC=4,2, RotorIO30401.iDestinationPos);(*4是左排，5是右排。左排转，右排不转*)
				MOV(ComConveyorIO30111.i_iResponsPCPLC=5,1, RotorIO30401.iDestinationPos);				
				IF (ComConveyorIO30111.i_iResponsPCPLC=4 AND  RotorIO30401.iCurrentPos=2 AND X61 )(*需要转，则等转到位置2,*)
					OR (ComConveyorIO30111.i_iResponsPCPLC=5 AND  RotorIO30401.iCurrentPos=1 AND X60 ) THEN(*不转则位置1为完成*)
					m_xRotor30401Done:=1;
				ELSE
						m_xRotor30401Done:=0;	
				END_IF;	
			ELSE(*无料就旋转回去，复位完成信号*)
				RotorIO30401.iDestinationPos:=1;
					m_xRotor30401Done:=0;
			END_IF;	
	(*预化成1入库转台下料*)		
	ConveyorIO30134.xUnload:=ConveyorIO30112.xEmpty 
														AND m_xRotor30401Done
														AND LifterIO30215.iCurrentPos=1 AND X5D;(*升降气缸*)
	ConveyorIO30112.xLoad:=ConveyorIO30134.xNextRun;
	IF ldp(TRUE,ConveyorIO30134.diDesConveyorOut>0) THEN
		ConveyorIO30112.diDesConveyorIn:=ConveyorIO30134.diDesConveyorOut;
		ConveyorIO30112.iTaskIDIn:=ConveyorIO30134.iTaskIDOut;
		ConveyorIO30112.iProductCategoryIn:=ConveyorIO30134.iProductCategoryOut;
	END_IF;
	(*预化成1入库气缸顶起*)
	LifterIO30215.xMDIExe:=NOT ConveyorIO30112.xError AND NOT ConveyorIO30112.xBusy;
	IF NOT ConveyorIO30112.xEmpty THEN
		LifterIO30215.iDestinationPos:=2;
	ELSE
		LifterIO30215.iDestinationPos:=1;
	END_IF;		
(***********************1巷道出库转台处理，运到转台上*********************)
	(*预化成1出库升降台控制*)
		IF ConveyorIO30114.xEmpty (*出库这里的开关位置要更改，改高点，不然putinto信号刷不到*)
			AND NOT ConveyorIO30114.xCWPresent
			AND NOT ConveyorIO30114.xCCWPresent
			AND NOT ConveyorIO30114.xBusy THEN
				LifterIO30214.iDestinationPos:=2;	
		ELSIF NOT ConveyorIO30114.xEmpty THEN
				LifterIO30214.iDestinationPos:=1;
		END_IF;	
			LifterIO30214.xMDIExe:=NOT ConveyorIO30114.xError AND NOT ConveyorIO30133.xError;
			DMOVP(ComConveyorIO30114.i_iResponsPCPLC=4,4,ConveyorIO30114.diDesConveyor);(*【需不需要转台转的信号生成】*)
			DMOVP(ComConveyorIO30114.i_iResponsPCPLC=5,5,ConveyorIO30114.diDesConveyor);(*【需不需要转台转的信号生成】*)			
			ConveyorIO30133.diDesConveyorIn:=ConveyorIO30114.diDesConveyorOut;(*【传递给转台】*)
			ConveyorIO30114.xUnload:=LifterIO30214.iCurrentPos=1 AND X5B(*升降台放下来*)
																	AND RotorIO30402.iCurrentPos=1 AND X62(*转台在接料位*)
																	 AND ConveyorIO30133.xEmpty(*转台为空*)
																	 AND ComConveyor30114.o_xReqSuccess(*旋转信号接收成功*);
			ConveyorIO30133.xLoad:=ConveyorIO30114.xNextRun;
	(*预化成1出库转台旋转控制*)		
		RotorIO30402.xMDIExe:=NOT ConveyorIO30133.xError AND NOT ConveyorIO30114.xError;
			IF NOT ConveyorIO30133.xEmpty THEN(*有料时，旋转，转到2旋转完成*)
				ConveyorIO30133.xUnloadCCW:=ConveyorIO30133.diDesConveyor=4;
				MOV(ConveyorIO30133.diDesConveyor=4,2, RotorIO30402.iDestinationPos);
				MOV(ConveyorIO30133.diDesConveyor=5,1, RotorIO30402.iDestinationPos);				
				IF (ConveyorIO30133.diDesConveyor=4 AND  RotorIO30402.iCurrentPos=2 AND X63 )(*需要转，则等转到位置2,*)
					OR (ConveyorIO30133.diDesConveyor=5 AND  RotorIO30402.iCurrentPos=1 AND X62 ) THEN(*不转则位置1为完成*)
					m_xRotor30402Done:=1;
				ELSE
					m_xRotor30402Done:=0;	
				END_IF;	
			ELSE(*无料就旋转回去，复位完成信号*)
				RotorIO30402.iDestinationPos:=1;
				m_xRotor30402Done:=0;
			END_IF;		
	(*化成1出库转台下料*)
		ConveyorIO30133.xUnload:=ConveyorIO30113.xEmpty 
														AND m_xRotor30402Done
														AND m_iTask30306=1;(*出库任务*)
(***********************1巷道出库的抢占任务，一边是产品出口，一边是2巷道的料路过*********************)	
	Task30306(xCondition:= Task30306Condition,
						xTaskComplete:= LDP(TRUE,ConveyorIO30110.xEmpty AND ConveyorIO30138.xEmpty ),
	 					xReset:=g_xResetSingle AND g_diDeviceIDSelect=30110,
						 iPriority:=m_iTask30306);
		Task30306Condition[1]:=NOT ConveyorIO30133.xEmpty AND  m_xRotor30402Done ;(*正常出库*)(*这里需要等待旋转完成信号*)
		Task30306Condition[2]:=NOT ConveyorIO30106.xEmpty AND  ConveyorIO30106.diDesConveyor=30116;(*2巷道的入库要料*)
	(*以上是1巷道出库顶升移载的抢占任务*)
	SwitchIO30306.xEntryEnable:=ConveyorIO30133.xNextRun;
	SwitchIO30306.xSwithEnable:=1;
	SwitchIO30306.xExitEnable:=ConveyorIO30138.xEmpty;
	(*任务2,去2巷道任务*)
	IF m_iTask30306=2 THEN
		IF ConveyorIO30110.xEmpty AND ConveyorIO30138.xEmpty THEN
			SwitchIO30306.xLiftCylinderExtend:=0;
			SwitchIO30306.xLiftCylinderRetract:=1;
		END_IF;
		ConveyorIO30110.xLoad:=ConveyorIO30106.xNextRun;
		ConveyorIO30110.diDesConveyorIn:=ConveyorIO30106.diDesConveyorOut;
		DMOVP(NOT ConveyorIO30110.xEmpty,ConveyorIO30106.diDesConveyor,ConveyorIO30113.diDesConveyor);(*【switch只能把目标地址传给入conveyor，不然会被写成0】*)
		SET(LDP(TRUE,NOT ConveyorIO30110.xEmpty),ConveyorIO30113.xPutInto);(*这里只要putinto了，就会进入switch正常流程了*)
		RST(LDP(TRUE,NOT ConveyorIO30113.xEmpty),ConveyorIO30113.xPutInto);	
	END_IF;
	(*任务为1时，顶升先升一下*)